VERSION : 0.1
   VAR_INPUT
      ix_SearchingMode : Bool;   // Searching button is pressed
      ix_EStop_Fbd : Bool;
      ix_LaserSensor : Bool;
   END_VAR
   VAR
      Available : Bool;   // At least sensor is available
      AxisControl : Array[0..2] of "UDT_AxisControl";
      AxisStatus : Array[0..2] of "UDT_AxisStatus";
      AxisX_Beginning : Bool;   // The X axis is in the start position
      AxisY_Beginning : Bool;   // The Y axis is in the start position
      AxisZ_Beginning : Bool;   // The Zaxis is in the start position
      StartBeginning : Bool;
      MoveY : Bool;
      ix_Enable : Bool;   // Search function is allowed
      Rtrig : Bool;
      SetCounter : Bool;   // Set the initial value of the state
   END_VAR
   VAR_TEMP
      "a" : Bool;
   END_VAR
   VAR_TEMP   // added for the SCL form of the ladder/FBD networks
      _w1 : Bool;
      _w2 : Bool;
   END_VAR
   // // AxisStatus[0] : X Axis
   // // AxisStatus[1] : Y Axis
   // // AxisStatus[2] : Z Axis
BEGIN

REGION Network 1: Search function is allowed
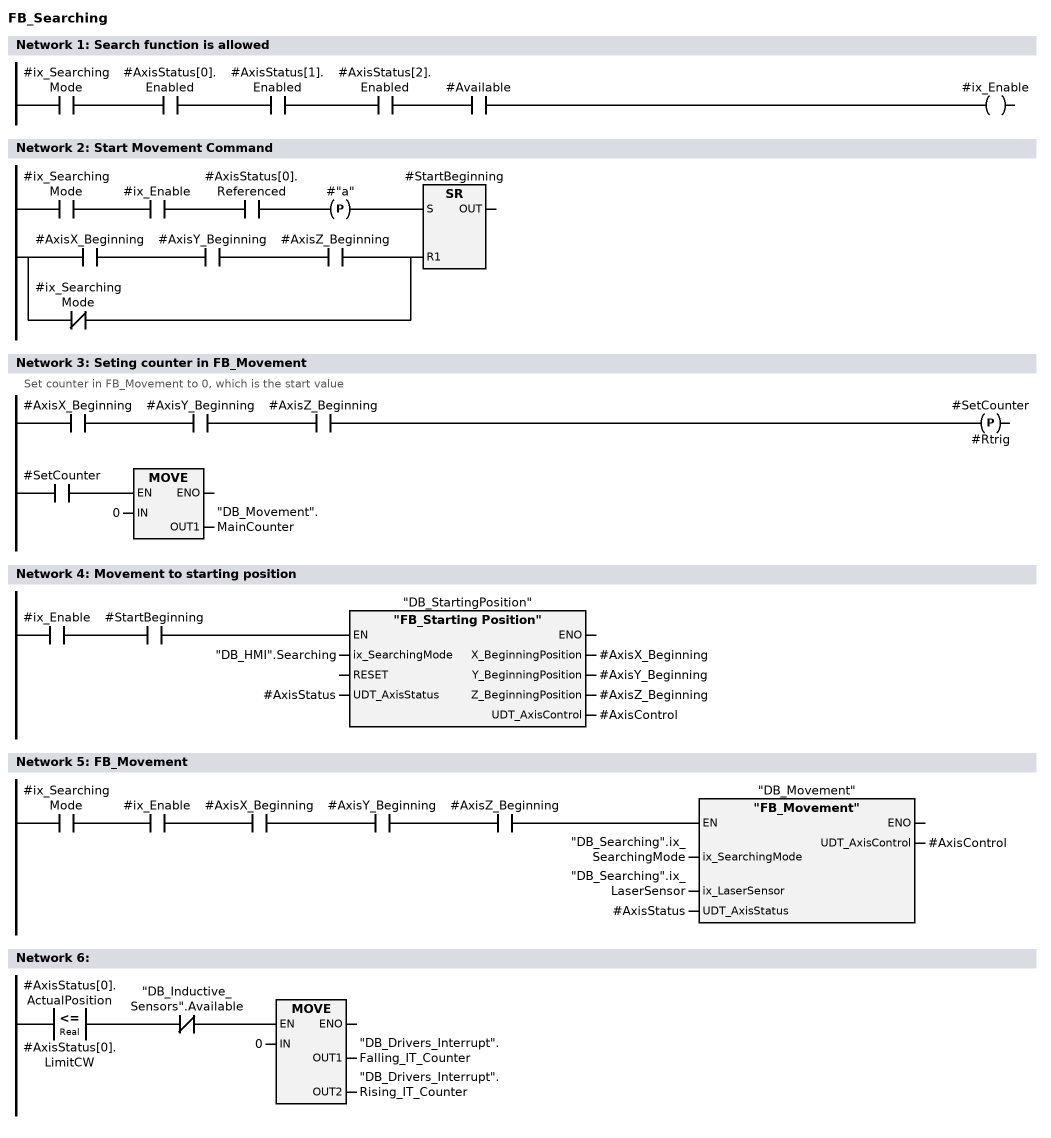
   RUNG wire#powerrail
      Contact( #ix_SearchingMode )
      Contact( #AxisStatus[0].Enabled )
      Contact( #AxisStatus[1].Enabled )
      Contact( #AxisStatus[2].Enabled )
      Contact( #Available )
      Coil( #ix_Enable )
   END_RUNG
   // the same network as SCL:
   #ix_Enable := #ix_SearchingMode AND #AxisStatus[0].Enabled AND #AxisStatus[1].Enabled AND #AxisStatus[2].Enabled AND #Available;
END_REGION

REGION Network 2: Start Movement Command
   RUNG wire#powerrail
      Contact( #ix_SearchingMode )
      Contact( #ix_Enable )
      Contact( #AxisStatus[0].Referenced )
      P_Trig( #"a" )
      S_SR(operand := #StartBeginning, r1 := wire#w1)
   END_RUNG
   RUNG wire#powerrail
      Contact( #AxisX_Beginning )
      Contact( #AxisY_Beginning )
      Contact( #AxisZ_Beginning )
   END_RUNG wire#w1
   RUNG wire#powerrail
      I_Contact( #ix_SearchingMode )
   END_RUNG wire#w1
   // the same network as SCL:
   #_w1 := #ix_SearchingMode AND #ix_Enable AND #AxisStatus[0].Referenced;
   #_w2 := #_w1 AND NOT #"a";   // rising edge
   #"a" := #_w1;
   IF #_w2 THEN
       #StartBeginning := TRUE;   // SR flip-flop
   END_IF;
   IF (#AxisX_Beginning AND #AxisY_Beginning AND #AxisZ_Beginning) OR NOT #ix_SearchingMode THEN
       #StartBeginning := FALSE;
   END_IF;
END_REGION

REGION Network 3: Seting counter in FB_Movement
   // Set counter in FB_Movement to 0, which is the start value
   #_w1 := #AxisX_Beginning AND #AxisY_Beginning AND #AxisZ_Beginning;
   #SetCounter := #_w1 AND NOT #Rtrig;   // rising edge
   #Rtrig := #_w1;
   IF #SetCounter THEN "DB_Movement".MainCounter := 0; END_IF;
END_REGION

REGION Network 4: Movement to starting position
   RUNG wire#powerrail
      Contact( #ix_Enable )
      Contact( #StartBeginning )
      "DB_StartingPosition"(ix_SearchingMode := "DB_HMI".Searching, RESET :=, UDT_AxisStatus := #AxisStatus, X_BeginningPosition => #AxisX_Beginning, Y_BeginningPosition => #AxisY_Beginning, Z_BeginningPosition => #AxisZ_Beginning, UDT_AxisControl => #AxisControl)
   END_RUNG
   // the same network as SCL:
   IF #ix_Enable AND #StartBeginning THEN
       "DB_StartingPosition"(ix_SearchingMode := "DB_HMI".Searching,   // "FB_Starting Position"
                             UDT_AxisStatus := #AxisStatus,
                             X_BeginningPosition => #AxisX_Beginning,
                             Y_BeginningPosition => #AxisY_Beginning,
                             Z_BeginningPosition => #AxisZ_Beginning,
                             UDT_AxisControl => #AxisControl);
   END_IF;
END_REGION

REGION Network 5: FB_Movement
   RUNG wire#powerrail
      Contact( #ix_SearchingMode )
      Contact( #ix_Enable )
      Contact( #AxisX_Beginning )
      Contact( #AxisY_Beginning )
      Contact( #AxisZ_Beginning )
      "DB_Movement"(ix_SearchingMode := "DB_Searching".ix_SearchingMode, ix_LaserSensor := "DB_Searching".ix_LaserSensor, UDT_AxisStatus := #AxisStatus, UDT_AxisControl => #AxisControl)
   END_RUNG
   // the same network as SCL:
   IF #ix_SearchingMode AND #ix_Enable AND #AxisX_Beginning AND #AxisY_Beginning AND #AxisZ_Beginning THEN
       "DB_Movement"(ix_SearchingMode := "DB_Searching".ix_SearchingMode,   // "FB_Movement"
                     ix_LaserSensor := "DB_Searching".ix_LaserSensor,
                     UDT_AxisStatus := #AxisStatus,
                     UDT_AxisControl => #AxisControl);
   END_IF;
END_REGION

REGION Network 6
   RUNG wire#powerrail
      { S7_Templates := "SrcType := Real" } LE_Contact(in1 := #AxisStatus[0].ActualPosition, in2 := #AxisStatus[0].LimitCW)
      I_Contact( "DB_Inductive_Sensors".Available )
      Move(in := 0, out1 => "DB_Drivers_Interrupt".Falling_IT_Counter, out2 => "DB_Drivers_Interrupt".Rising_IT_Counter)
   END_RUNG
   // the same network as SCL:
   IF (#AxisStatus[0].ActualPosition <= #AxisStatus[0].LimitCW) AND NOT "DB_Inductive_Sensors".Available THEN
       "DB_Drivers_Interrupt".Falling_IT_Counter := 0;
       "DB_Drivers_Interrupt".Rising_IT_Counter := 0;
   END_IF;
END_REGION
END_FUNCTION_BLOCK

// folder: Searching Mode/Movement

FUNCTION_BLOCK "FB_Movement"   // FB4, LAD
{ S7_Optimized_Access := 'TRUE' }
VERSION : 0.1
   VAR_INPUT
      ix_SearchingMode : Bool;
      ix_LaserSensor : Bool;
      UDT_AxisStatus : Array[0..2] of "UDT_AxisStatus";
   END_VAR
   VAR_OUTPUT
      UDT_AxisControl : Array[0..2] of "UDT_AxisControl";
   END_VAR
   VAR
      MainCounter : Int;   // Main counter show which part of the code is performing in this moment
      YAxisLimit : Real := 20.0;   // Min limit of the Y Axis
      NewYPos : Real;   // New Y required position
      Ymin : Int;
      Ymax : Int;
      RTrigCount0 : Bool;
      Reset1 : Bool;
      PTrigCount2 : Bool;
      Reset2 : Bool;
      Start : Struct
         X : Struct
            Right : Array[0..1] of Bool;
            Left : Array[0..1] of Bool;
            "Repeat" : Bool;
         END_STRUCT;
         Y : Array[0..3] of Bool;
         ReturnToStartPos : Bool;
         RepeatY : Bool;
      END_STRUCT;
      Ptrig : Struct
         X : Struct
            Right : Array[0..1] of Bool;
            Left : Array[0..1] of Bool;
            "Repeat" : Bool;
         END_STRUCT;
         Y : Array[0..3] of Bool;
         ReturnToStartPos : Bool;
      END_STRUCT;
      "Timer" : Array[0..2] of Bool;
   END_VAR
   VAR_TEMP   // added for the SCL form of the ladder/FBD networks
      _w1 : Bool;
      _w2 : Bool;
   END_VAR
BEGIN

REGION Network 1: General Counter
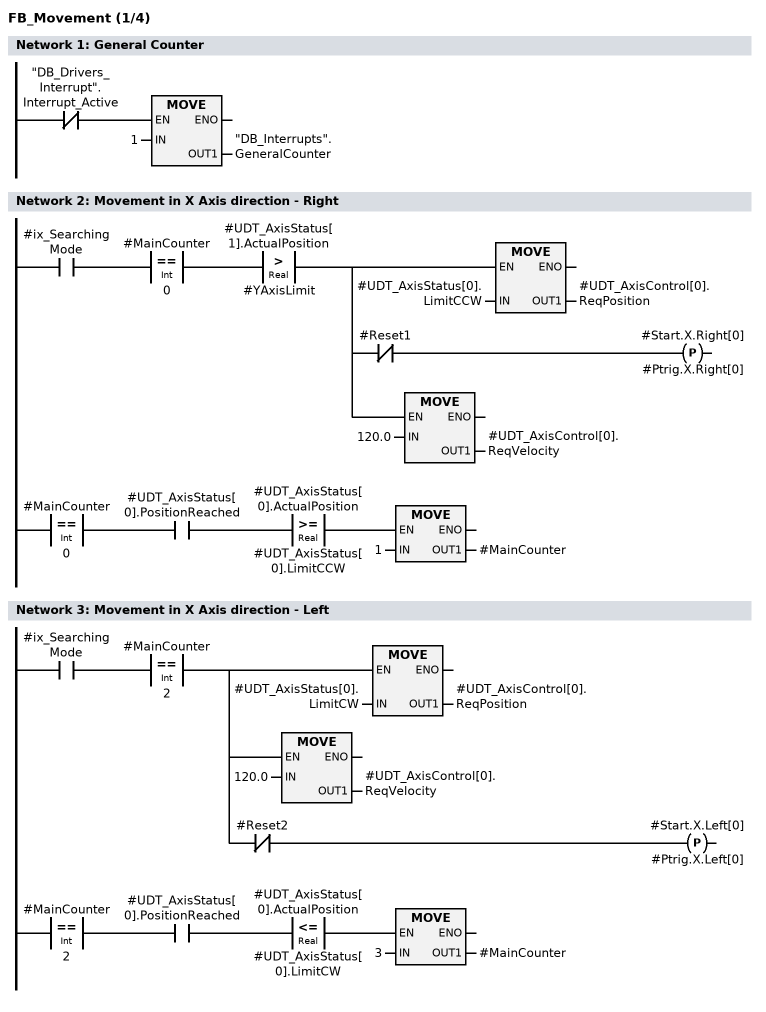
   RUNG wire#powerrail
      I_Contact( "DB_Drivers_Interrupt".Interrupt_Active )
      Move(in := 1, out1 => "DB_Interrupts".GeneralCounter)
   END_RUNG
   // the same network as SCL:
   IF NOT "DB_Drivers_Interrupt".Interrupt_Active THEN "DB_Interrupts".GeneralCounter := 1; END_IF;
END_REGION

REGION Network 2: Movement in X Axis direction - Right
   #_w1 := #ix_SearchingMode AND (#MainCounter = 0) AND (#UDT_AxisStatus[1].ActualPosition > #YAxisLimit);
   IF #_w1 THEN #UDT_AxisControl[0].ReqPosition := #UDT_AxisStatus[0].LimitCCW; END_IF;
   #_w2 := #_w1 AND NOT #Reset1;
   #Start.X.Right[0] := #_w2 AND NOT #Ptrig.X.Right[0];   // rising edge
   #Ptrig.X.Right[0] := #_w2;
   IF #_w1 THEN #UDT_AxisControl[0].ReqVelocity := 120.0; END_IF;
   IF (#MainCounter = 0) AND #UDT_AxisStatus[0].PositionReached AND (#UDT_AxisStatus[0].ActualPosition >= #UDT_AxisStatus[0].LimitCCW) THEN
       #MainCounter := 1;
   END_IF;
END_REGION

REGION Network 3: Movement in X Axis direction - Left
   #_w1 := #ix_SearchingMode AND (#MainCounter = 2);
   IF #_w1 THEN
       #UDT_AxisControl[0].ReqPosition := #UDT_AxisStatus[0].LimitCW;
       #UDT_AxisControl[0].ReqVelocity := 120.0;
   END_IF;
   #_w2 := #_w1 AND NOT #Reset2;
   #Start.X.Left[0] := #_w2 AND NOT #Ptrig.X.Left[0];   // rising edge
   #Ptrig.X.Left[0] := #_w2;
   IF (#MainCounter = 2) AND #UDT_AxisStatus[0].PositionReached AND (#UDT_AxisStatus[0].ActualPosition <= #UDT_AxisStatus[0].LimitCW) THEN
       #MainCounter := 3;
   END_IF;
END_REGION

REGION Network 4: Movement in Y axis
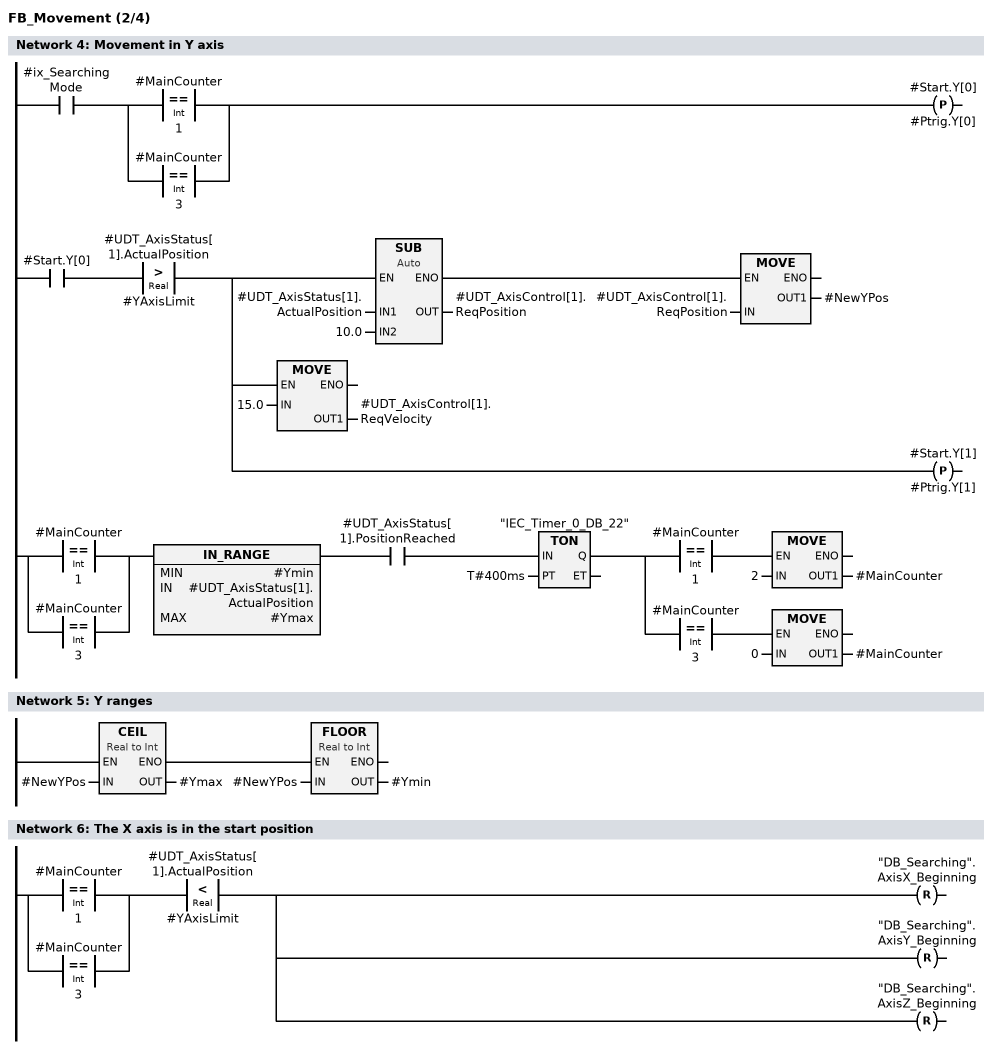
   #_w1 := #ix_SearchingMode AND ((#MainCounter = 1) OR (#MainCounter = 3));
   #Start.Y[0] := #_w1 AND NOT #Ptrig.Y[0];   // rising edge
   #Ptrig.Y[0] := #_w1;
   #_w2 := #Start.Y[0] AND (#UDT_AxisStatus[1].ActualPosition > #YAxisLimit);
   IF #_w2 THEN
       #UDT_AxisControl[1].ReqPosition := #UDT_AxisStatus[1].ActualPosition - 10.0;
       #NewYPos := #UDT_AxisControl[1].ReqPosition;
       #UDT_AxisControl[1].ReqVelocity := 15.0;
   END_IF;
   #Start.Y[1] := #_w2 AND NOT #Ptrig.Y[1];   // rising edge
   #Ptrig.Y[1] := #_w2;
   "IEC_Timer_0_DB_22".TON(IN := ((#MainCounter = 1) OR (#MainCounter = 3)) AND (#Ymin <= #UDT_AxisStatus[1].ActualPosition) AND (#UDT_AxisStatus[1].ActualPosition <= #Ymax) AND #UDT_AxisStatus[1].PositionReached,
                           PT := T#400ms);
   IF "IEC_Timer_0_DB_22".Q AND (#MainCounter = 1) THEN #MainCounter := 2; END_IF;
   IF "IEC_Timer_0_DB_22".Q AND (#MainCounter = 3) THEN #MainCounter := 0; END_IF;
END_REGION

REGION Network 5: Y ranges
   #Ymax := CEIL(#NewYPos);
   #Ymin := FLOOR(#NewYPos);
END_REGION

REGION Network 6: The X axis is in the start position
   RUNG wire#powerrail
      { S7_Templates := "SrcType := Int" } EQ_Contact(in1 := #MainCounter, in2 := 1)
      wire#w1
      { S7_Templates := "SrcType := Real" } LT_Contact(in1 := #UDT_AxisStatus[1].ActualPosition, in2 := #YAxisLimit)
      wire#w2
      R_Coil( "DB_Searching".AxisX_Beginning )
   END_RUNG
   RUNG wire#powerrail
      { S7_Templates := "SrcType := Int" } EQ_Contact(in1 := #MainCounter, in2 := 3)
   END_RUNG wire#w1
   RUNG wire#w2
      R_Coil( "DB_Searching".AxisY_Beginning )
   END_RUNG
   RUNG wire#w2
      R_Coil( "DB_Searching".AxisZ_Beginning )
   END_RUNG
   // the same network as SCL:
   IF ((#MainCounter = 1) OR (#MainCounter = 3)) AND (#UDT_AxisStatus[1].ActualPosition < #YAxisLimit) THEN
       "DB_Searching".AxisX_Beginning := FALSE;
       "DB_Searching".AxisY_Beginning := FALSE;
       "DB_Searching".AxisZ_Beginning := FALSE;
   END_IF;
END_REGION

REGION Network 7: Return from the interrupt
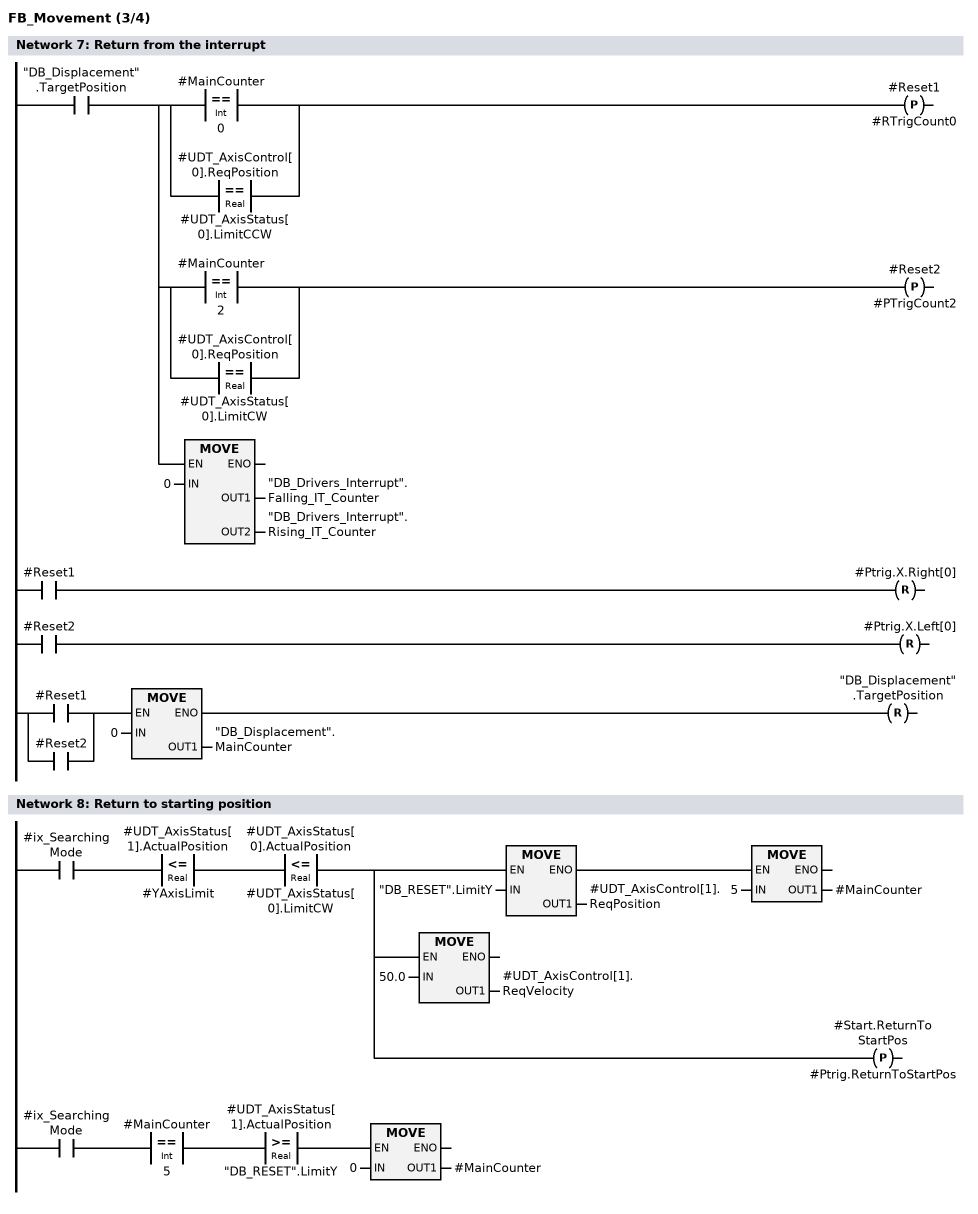
   #_w1 := "DB_Displacement".TargetPosition AND ((#MainCounter = 0) OR (#UDT_AxisControl[0].ReqPosition = #UDT_AxisStatus[0].LimitCCW));
   #Reset1 := #_w1 AND NOT #RTrigCount0;   // rising edge
   #RTrigCount0 := #_w1;
   #_w2 := "DB_Displacement".TargetPosition AND ((#MainCounter = 2) OR (#UDT_AxisControl[0].ReqPosition = #UDT_AxisStatus[0].LimitCW));
   #Reset2 := #_w2 AND NOT #PTrigCount2;   // rising edge
   #PTrigCount2 := #_w2;
   IF "DB_Displacement".TargetPosition THEN
       "DB_Drivers_Interrupt".Falling_IT_Counter := 0;
       "DB_Drivers_Interrupt".Rising_IT_Counter := 0;
   END_IF;
   IF #Reset1 THEN #Ptrig.X.Right[0] := FALSE; END_IF;
   IF #Reset2 THEN #Ptrig.X.Left[0] := FALSE; END_IF;
   IF #Reset1 OR #Reset2 THEN
       "DB_Displacement".MainCounter := 0;
       "DB_Displacement".TargetPosition := FALSE;
   END_IF;
END_REGION

REGION Network 8: Return to starting position
   #_w1 := #ix_SearchingMode AND (#UDT_AxisStatus[1].ActualPosition <= #YAxisLimit) AND (#UDT_AxisStatus[0].ActualPosition <= #UDT_AxisStatus[0].LimitCW);
   IF #_w1 THEN
       #UDT_AxisControl[1].ReqPosition := "DB_RESET".LimitY;
       #MainCounter := 5;
       #UDT_AxisControl[1].ReqVelocity := 50.0;
   END_IF;
   #Start.ReturnToStartPos := #_w1 AND NOT #Ptrig.ReturnToStartPos;   // rising edge
   #Ptrig.ReturnToStartPos := #_w1;
   IF #ix_SearchingMode AND (#MainCounter = 5) AND (#UDT_AxisStatus[1].ActualPosition >= "DB_RESET".LimitY) THEN
       #MainCounter := 0;
   END_IF;
END_REGION

REGION Network 9: Repeat pulse X Axis
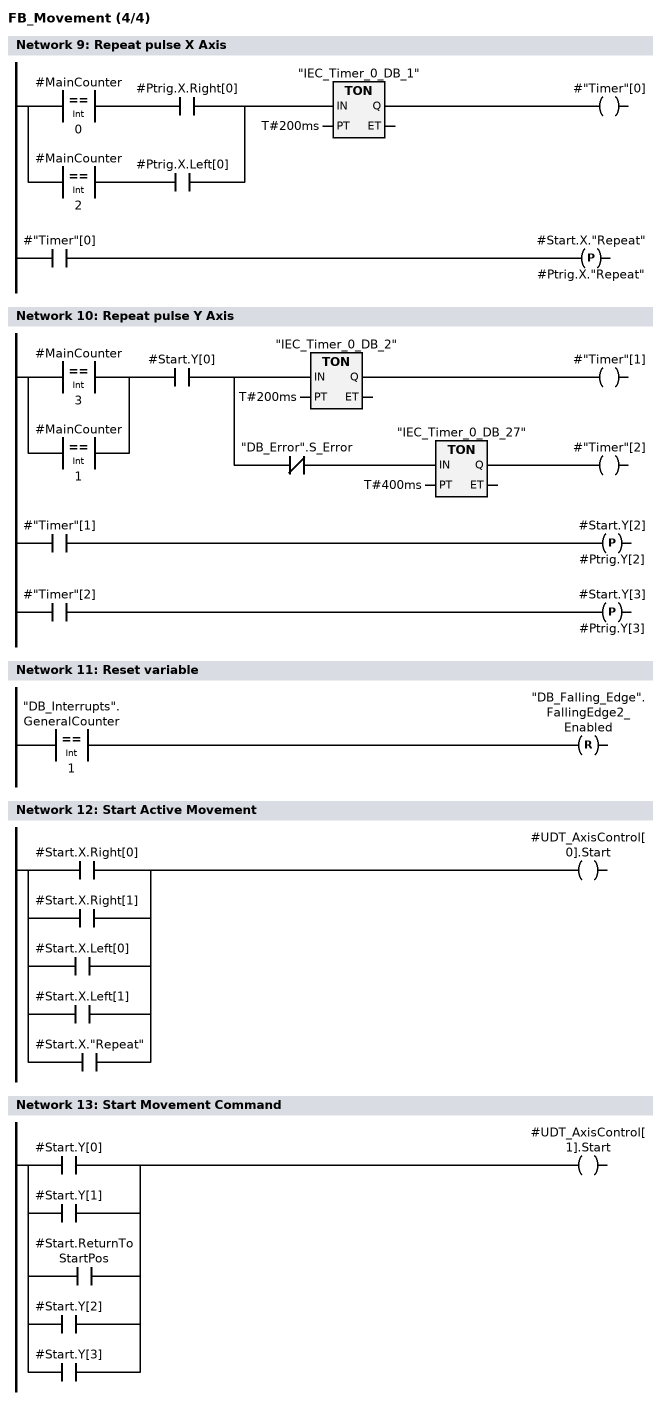
   "IEC_Timer_0_DB_1".TON(IN := ((#MainCounter = 0) AND #Ptrig.X.Right[0]) OR ((#MainCounter = 2) AND #Ptrig.X.Left[0]),
                          PT := T#200ms);
   #"Timer"[0] := "IEC_Timer_0_DB_1".Q;
   #Start.X."Repeat" := #"Timer"[0] AND NOT #Ptrig.X."Repeat";   // rising edge
   #Ptrig.X."Repeat" := #"Timer"[0];
END_REGION

REGION Network 10: Repeat pulse Y Axis
   #_w1 := ((#MainCounter = 3) OR (#MainCounter = 1)) AND #Start.Y[0];
   "IEC_Timer_0_DB_2".TON(IN := #_w1, PT := T#200ms);
   #"Timer"[1] := "IEC_Timer_0_DB_2".Q;
   "IEC_Timer_0_DB_27".TON(IN := #_w1 AND NOT "DB_Error".S_Error, PT := T#400ms);
   #"Timer"[2] := "IEC_Timer_0_DB_27".Q;
   #Start.Y[2] := #"Timer"[1] AND NOT #Ptrig.Y[2];   // rising edge
   #Ptrig.Y[2] := #"Timer"[1];
   #Start.Y[3] := #"Timer"[2] AND NOT #Ptrig.Y[3];   // rising edge
   #Ptrig.Y[3] := #"Timer"[2];
END_REGION

REGION Network 11: Reset variable
   RUNG wire#powerrail
      { S7_Templates := "SrcType := Int" } EQ_Contact(in1 := "DB_Interrupts".GeneralCounter, in2 := 1)
      R_Coil( "DB_Falling_Edge".FallingEdge2_Enabled )
   END_RUNG
   // the same network as SCL:
   IF "DB_Interrupts".GeneralCounter = 1 THEN "DB_Falling_Edge".FallingEdge2_Enabled := FALSE; END_IF;
END_REGION

REGION Network 12: Start Active Movement
   RUNG wire#powerrail
      Contact( #Start.X.Right[0] )
      wire#w1
      Coil( #UDT_AxisControl[0].Start )
   END_RUNG
   RUNG wire#powerrail
      Contact( #Start.X.Right[1] )
   END_RUNG wire#w1
   RUNG wire#powerrail
      Contact( #Start.X.Left[0] )
   END_RUNG wire#w1
   RUNG wire#powerrail
      Contact( #Start.X.Left[1] )
   END_RUNG wire#w1
   RUNG wire#powerrail
      Contact( #Start.X."Repeat" )
   END_RUNG wire#w1
   // the same network as SCL:
   #UDT_AxisControl[0].Start := #Start.X.Right[0] OR #Start.X.Right[1] OR #Start.X.Left[0] OR #Start.X.Left[1] OR #Start.X."Repeat";
END_REGION

REGION Network 13: Start Movement Command
   RUNG wire#powerrail
      Contact( #Start.Y[0] )
      wire#w1
      Coil( #UDT_AxisControl[1].Start )
   END_RUNG
   RUNG wire#powerrail
      Contact( #Start.Y[1] )
   END_RUNG wire#w1
   RUNG wire#powerrail
      Contact( #Start.ReturnToStartPos )
   END_RUNG wire#w1
   RUNG wire#powerrail
      Contact( #Start.Y[2] )
   END_RUNG wire#w1
   RUNG wire#powerrail
      Contact( #Start.Y[3] )
   END_RUNG wire#w1
   // the same network as SCL:
   #UDT_AxisControl[1].Start := #Start.Y[0] OR #Start.Y[1] OR #Start.ReturnToStartPos OR #Start.Y[2] OR #Start.Y[3];
END_REGION
END_FUNCTION_BLOCK

// folder: Searching Mode/Starting Position

FUNCTION_BLOCK "FB_Starting Position"   // FB5, LAD
{ S7_Optimized_Access := 'TRUE' }
VERSION : 0.1
   VAR_INPUT
      ix_SearchingMode : Bool;
      RESET : Bool;
      UDT_AxisStatus : Array[0..2] of "UDT_AxisStatus";
   END_VAR
   VAR_OUTPUT
      X_BeginningPosition : Bool;
      Y_BeginningPosition : Bool;
      Z_BeginningPosition : Bool;
      UDT_AxisControl : Array[0..2] of "UDT_AxisControl";
   END_VAR
   VAR
      Starting : Bool;
      RTrig : Bool;
      Start : Bool;
      LIMITY : Real;
   END_VAR
BEGIN

REGION Network 1
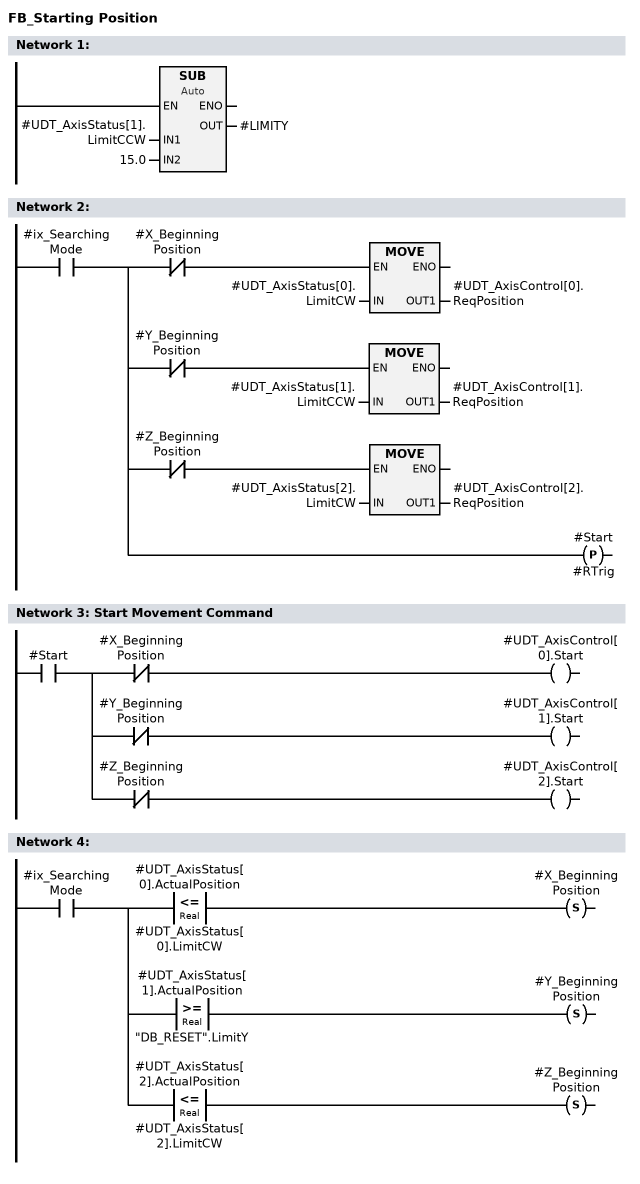
   RUNG wire#powerrail
      Sub(in1 := #UDT_AxisStatus[1].LimitCCW, in2 := 15.0, out => #LIMITY)
   END_RUNG
   // the same network as SCL:
   #LIMITY := #UDT_AxisStatus[1].LimitCCW - 15.0;
END_REGION

REGION Network 2
   IF #ix_SearchingMode AND NOT #X_BeginningPosition THEN
       #UDT_AxisControl[0].ReqPosition := #UDT_AxisStatus[0].LimitCW;
   END_IF;
   IF #ix_SearchingMode AND NOT #Y_BeginningPosition THEN
       #UDT_AxisControl[1].ReqPosition := #UDT_AxisStatus[1].LimitCCW;
   END_IF;
   IF #ix_SearchingMode AND NOT #Z_BeginningPosition THEN
       #UDT_AxisControl[2].ReqPosition := #UDT_AxisStatus[2].LimitCW;
   END_IF;
   #Start := #ix_SearchingMode AND NOT #RTrig;   // rising edge
   #RTrig := #ix_SearchingMode;
END_REGION

REGION Network 3: Start Movement Command
   RUNG wire#powerrail
      Contact( #Start )
      wire#w1
      I_Contact( #X_BeginningPosition )
      Coil( #UDT_AxisControl[0].Start )
   END_RUNG
   RUNG wire#w1
      I_Contact( #Y_BeginningPosition )
      Coil( #UDT_AxisControl[1].Start )
   END_RUNG
   RUNG wire#w1
      I_Contact( #Z_BeginningPosition )
      Coil( #UDT_AxisControl[2].Start )
   END_RUNG
   // the same network as SCL:
   #UDT_AxisControl[0].Start := #Start AND NOT #X_BeginningPosition;
   #UDT_AxisControl[1].Start := #Start AND NOT #Y_BeginningPosition;
   #UDT_AxisControl[2].Start := #Start AND NOT #Z_BeginningPosition;
END_REGION

REGION Network 4
   RUNG wire#powerrail
      Contact( #ix_SearchingMode )
      wire#w1
      { S7_Templates := "SrcType := Real" } LE_Contact(in1 := #UDT_AxisStatus[0].ActualPosition, in2 := #UDT_AxisStatus[0].LimitCW)
      S_Coil( #X_BeginningPosition )
   END_RUNG
   RUNG wire#w1
      { S7_Templates := "SrcType := Real" } GE_Contact(in1 := #UDT_AxisStatus[1].ActualPosition, in2 := "DB_RESET".LimitY)
      S_Coil( #Y_BeginningPosition )
   END_RUNG
   RUNG wire#w1
      { S7_Templates := "SrcType := Real" } LE_Contact(in1 := #UDT_AxisStatus[2].ActualPosition, in2 := #UDT_AxisStatus[2].LimitCW)
      S_Coil( #Z_BeginningPosition )
   END_RUNG
   // the same network as SCL:
   IF #ix_SearchingMode AND (#UDT_AxisStatus[0].ActualPosition <= #UDT_AxisStatus[0].LimitCW) THEN
       #X_BeginningPosition := TRUE;
   END_IF;
   IF #ix_SearchingMode AND (#UDT_AxisStatus[1].ActualPosition >= "DB_RESET".LimitY) THEN
       #Y_BeginningPosition := TRUE;
   END_IF;
   IF #ix_SearchingMode AND (#UDT_AxisStatus[2].ActualPosition <= #UDT_AxisStatus[2].LimitCW) THEN
       #Z_BeginningPosition := TRUE;
   END_IF;
END_REGION
END_FUNCTION_BLOCK

(* ===== HMI "HMI_RT" =====
system functions are stored by id; their names below are inferred from use
connection "HMI_Connection": ETHERNET, SMART_S7_1200_OMS

HMI tags "Default tag table"
   "DB_HMI_Reset" : Bool = PLC DB_HMI.Reset AT %DB1.DBW0, 500 ms
   "DB_HMI_Enable" : Bool = PLC DB_HMI.Enable AT %DB1.DBX0.0, 500 ms
   "ScreenNumber" : Int AT %DB1.DBW0
   "EStop_Fdb" : Bool = PLC EStop_Fdb AT %I8.6, 500 ms
   "DB_HMI_Searching" : Bool = PLC DB_HMI.Searching, 1 s
   "DB_HMI_StartPosition" : Bool = PLC DB_HMI.StartPosition, 1 s
   "DB_HMI_Interrupt" : Bool = PLC DB_HMI.Interrupt, 100 ms
   "DB_HMI_Electromagnet" : Bool = PLC DB_HMI.Electromagnet, 500 ms
   "Laser Sensor" : Bool = PLC "Laser Sensor" AT %I0.0, 1 s
   "Drivers_DB_UDT_Axis_Status{0}_LimitCW" : Real = PLC DB_Drivers.UDT_Axis_Status[0].LimitCW, 1 s
   "Drivers_DB_UDT_Axis_Status{0}_ActualPosition" : Real = PLC DB_Drivers.UDT_Axis_Status[0].ActualPosition, 100 ms
   "Drivers_DB_UDT_Axis_Status{0}_ActualVelocity" : Real = PLC DB_Drivers.UDT_Axis_Status[0].ActualVelocity, 100 ms
   "Drivers_DB_UDT_Axis_Status{0}_LimitCCW" : Real = PLC DB_Drivers.UDT_Axis_Status[0].LimitCCW, 1 s
   "FB_Axis_Y_DB_o_Status_ActualPosition" : Real = PLC FB_Axis_Y_DB.o_Status.ActualPosition, 100 ms
   "FB_Axis_Y_DB_o_Status_ActualVelocity" : Real = PLC FB_Axis_Y_DB.o_Status.ActualVelocity, 100 ms
   "FB_Axis_Y_DB_o_Status_LimitCW" : Real = PLC FB_Axis_Y_DB.o_Status.LimitCW, 1 s
   "FB_Axis_Y_DB_o_Status_LimitCCW" : Real = PLC FB_Axis_Y_DB.o_Status.LimitCCW, 1 s
   "FB_Axis_Z_DB_o_Status_ActualPosition" : Real = PLC FB_Axis_Z_DB.o_Status.ActualPosition, 100 ms
   "FB_Axis_Z_DB_o_Status_ActualVelocity" : Real = PLC FB_Axis_Z_DB.o_Status.ActualVelocity, 100 ms
   "FB_Axis_Z_DB_o_Status_LimitCW" : Real = PLC FB_Axis_Z_DB.o_Status.LimitCW, 1 s
   "FB_Axis_Z_DB_o_Status_LimitCCW" : Real = PLC FB_Axis_Z_DB.o_Status.LimitCCW, 1 s
   "FB_Axis_Z_DB_o_Status_Error" : Bool = PLC FB_Axis_Z_DB.o_Status.Error, 1 s
   "FB_Axis_Y_DB_o_Status_Error" : Bool = PLC FB_Axis_Y_DB.o_Status.Error, 1 s
   "FB_Axis_X_DB_o_Status_Error" : Bool = PLC FB_Axis_X_DB.o_Status.Error, 1 s
   "Interrupts_DB_GeneralCounter" : Int = PLC DB_Interrupts.GeneralCounter, 100 ms
   "FallingEdge_DB_Enabled" : Bool = PLC DB_Falling_Edge.Enabled, 1 s
   "FallingEdge2_DB_Enabled" : Bool = PLC DB_Line2.Enabled, 1 s
   "Drivers_DB_X_AVG" : Real = PLC DB_Drivers.X_AVG, 1 s
   "Drivers_DB_Y_AVG" : Real = PLC DB_Drivers.Y_AVG, 1 s
   "Drivers_Interrupt_DB_Interrupt_Active" : Bool = PLC DB_Drivers_Interrupt.Interrupt_Active, 1 s
   "DB_HMI_AvailablePlace" : Int = PLC DB_HMI.AvailablePlace, 100 ms
   "DB_HMI_Error" : Bool = PLC DB_HMI.Error, 100 ms
   "DB_HMI_Start/Enable" : Bool = PLC DB_HMI.Start/Enable, 100 ms
   "DB_HMI_MidPosCounting" : Bool = PLC DB_HMI.MidPosCounting, 100 ms
   "DB_HMI_ItemwasFound" : Bool = PLC DB_HMI.ItemwasFound, 100 ms
   "DB_HMI_GrabbingTheItem" : Bool = PLC DB_HMI.GrabbingTheItem, 100 ms
   "DB_HMI_StartPositionReached" : Bool = PLC DB_HMI.StartPositionReached, 100 ms
   "DB_HMI_MovingToStartPosition" : Bool = PLC DB_HMI.MovingToStartPosition, 100 ms
   "DB_HMI_ErrorState" : Int = PLC DB_HMI.ErrorState, 500 ms
   "DB_HMI_ResetError" : Bool = PLC DB_HMI.ResetError, 500 ms
   "DB_HMI_ResetSpace" : Bool = PLC DB_HMI.ResetSpace, 1 s
   "DB_HMI_PlaceOcc_S1" : Bool = PLC DB_HMI.PlaceOcc.S1, 1 s
   "DB_HMI_PlaceOcc_S2" : Bool = PLC DB_HMI.PlaceOcc.S2, 1 s
   "DB_HMI_PlaceOcc_S3" : Bool = PLC DB_HMI.PlaceOcc.S3, 1 s
   "DB_HMI_PlaceOcc_S4" : Bool = PLC DB_HMI.PlaceOcc.S4, 1 s
   "DB_Displacement_PlaceOcup_Sens1" : Bool = PLC DB_Displacement.PlaceOcup.Sens1, 1 s
   "DB_Displacement_PlaceOcup_Sens2" : Bool = PLC DB_Displacement.PlaceOcup.Sens2, 1 s
   "DB_Displacement_PlaceOcup_Sens3" : Bool = PLC DB_Displacement.PlaceOcup.Sens3, 1 s
   "DB_Displacement_PlaceOcup_Sens4" : Bool = PLC DB_Displacement.PlaceOcup.Sens4, 1 s